
           // -------------------------------------------------------
       10: // Esperar a que el KRC pida número de programa (PGNO_REQ = 1)
           IF #ROB_PGNO_REQ THEN
               // Latch del programa seleccionado (1..3). Forzamos límites por seguridad.
               IF #ProgSel < USINT#1 THEN
                   #pgnoLatched := USINT#1;
               ELSIF #ProgSel > USINT#3 THEN
                   #pgnoLatched := USINT#3;
               ELSE
                   #pgnoLatched := #ProgSel;
               END_IF;

               #step := 20;
           END_IF;


       20: // Presentar PGNO MIENTRAS PGNO_REQ = 1
           IF #ROB_PGNO_REQ THEN
               // Escribir bits binarios 101..108 a partir de #pgnoLatched
               #PGNO_101 := ((#pgnoLatched AND USINT#1) <> USINT#0);
               #PGNO_102 := ((#pgnoLatched AND USINT#2) <> USINT#0);
               #PGNO_103 := ((#pgnoLatched AND USINT#4) <> USINT#0);
               #PGNO_104 := ((#pgnoLatched AND USINT#8) <> USINT#0);
               #PGNO_105 := ((#pgnoLatched AND USINT#16) <> USINT#0);
               #PGNO_106 := ((#pgnoLatched AND USINT#32) <> USINT#0);
               #PGNO_107 := ((#pgnoLatched AND USINT#64) <> USINT#0);
               #PGNO_108 := ((#pgnoLatched AND USINT#128) <> USINT#0);

               // Paridad "even": XOR de los 8 bits (1 si nº de unos es impar)
               #PGNO_PARITY :=
               #PGNO_101 XOR #PGNO_102 XOR #PGNO_103 XOR #PGNO_104 XOR
               #PGNO_105 XOR #PGNO_106 XOR #PGNO_107 XOR #PGNO_108;

               // Arrancamos el TON de estabilidad y pasamos a validación
               #tStable(IN := TRUE,
                        PT := #stableTime);
               #step := 21;
           END_IF;


       21: // Esperar estabilidad y marcar PGNO_VALID
           #tStable(IN := (#step = 21),
                    PT := #stableTime);
           IF #tStable.Q THEN
               #PGNO_VALID := TRUE;        // el KRC ya puede muestrear PGNO
               #step := 22;
           END_IF;


       22: // Mantener PGNO_VALID hasta la CAÍDA de PGNO_REQ
           #PGNO_VALID := TRUE;
           IF #fPgnoReq.Q THEN
               #PGNO_VALID := FALSE;    // cerrar handshake de selección

               // limpiar PGNO para siguientes ciclos
               #PGNO_101 := FALSE;
               #PGNO_102 := FALSE;
               #PGNO_103 := FALSE;
               #PGNO_104 := FALSE;
               #PGNO_105 := FALSE;
               #PGNO_106 := FALSE;
               #PGNO_107 := FALSE;
               #PGNO_108 := FALSE;
               #PGNO_PARITY := FALSE;

               #step := 40;    // → arranque real del programa
           END_IF;

       40: // START real: segundo pulso de $EXT_START para ejecutar el programa
           "ALM_FILTER" := TRUE; // marcador/diagnóstico ELIMINAR
           #tpStart(IN := TRUE,
                    PT := #pulseTime);
           #EXT_START := #tpStart.Q;
           IF NOT #tpStart.Q THEN
               #ROBOT_READY := TRUE;   // handshake completo
               #step := 60;            // → ejecución
           END_IF;


       60: // En ejecución / rearme
           // Para un nuevo ciclo hay que hacer hacer 0→1 de nuevo desde la aplicacion 
           // si #startAutExt no baja, #rStart.Q no volverá a disparar.
           #step := 0;

   END_CASE;
END_REGION
END_FUNCTION_BLOCK

// folder: 20. Robot Services/Mov Manual

FUNCTION_BLOCK "TcpJogging"   // FB5, LAD
{ S7_Optimized_Access := 'TRUE' }
VERSION : 0.1
   VAR_INPUT
      "buttonX+" : Bool;
      "buttonX-" : Bool;
      "buttonY+" : Bool;
      "buttonY-" : Bool;
      "buttonZ+" : Bool;
      "buttonZ-" : Bool;
      "buttonE1+" : Bool;
      "buttonE1-" : Bool;
   END_VAR
BEGIN

REGION Network 1 (SCL): Mapea los valores de los botones de WF
   IF "PlcStatus".mode.effective = 0 THEN

       "Tag_1" := TRUE;
       //MOV X,Y,Z
       //%Q630.0 = buttonX+
       //%Q630.1 = buttonX-
       //%Q630.2 = buttonY+
       //%Q630.3 = buttonY-
       //%Q630.4 = buttonZ+
       //%Q630.5 = buttonZ-
       //MOV A,B,C
       //%Q630.6 = buttonWF +A
       //%Q630.7 = buttonWF -A
       //%Q631.0 = buttonWF +B
       //%Q631.1 = buttonWF -B
       //%Q631.2 = buttonWF +C
       //%Q631.3 = buttonWF -C
       //Mov E1
       //%Q631.4 = buttonWF +E1
       //%Q631.5 = buttonWF -E1

   ELSE
       //%Q631.1 = buttonWF -B
       "Tag_1" := FALSE;
   END_IF;
END_REGION
END_FUNCTION_BLOCK

FUNCTION_BLOCK "TcpTarget"   // FB11, LAD
{ S7_Optimized_Access := 'TRUE' }
VERSION : 0.1
   VAR_INPUT
      KukaControlCmdCode : UInt;
      KukaControlCmdSeq : UInt;
      KukaControlCmdProfileRequestId : UInt;
      KukaControlCmdToolRequestId : UInt;
      KukaControlCmdBaseRequestId : UInt;
      KukaControlCmdProgramRequestId : UInt;
      KukaControlTcpTargetX_mm : LReal;
      KukaControlTcpTargetY_mm : LReal;
      KukaControlTcpTargetZ_mm : LReal;
      kukaControlE1Target_mm : LReal;
      KukaControlCmdCancelGo : Bool;
      KukaControlCmdPauseGo : Bool;
      KukaControlCmdResumeGo : Bool;
      enterService : Bool;
      KukaControlCmdVel : UInt;
      KukaControlCmdIndex : UInt;
      scanPuntoInicialX : LReal;
      scanPuntoInicialY : LReal;
      scanPuntoInicialZ : LReal;
      scanPuntoInicialE1 : LReal;
      scanPuntoFinalX : LReal;
      scanPuntoFinalY : LReal;
      scanPuntoFinalZ : LReal;
      scanPuntoFinalE1 : LReal;
   END_VAR
   VAR_OUTPUT
      moveCodeKuka : Word;
      profileReqId : Word;
      baseReqId : Word;
      toolReqId : Word;
      programReqId : Word;
      x_mmHe : DWord;
      y_mmHe : DWord;
      z_mmHe : DWord;
      e_mmHe : DWord;
      PlcStatusExecDone : Bool;
      PlcStatusExecAccepted : Bool;
      PlcStatusExecAckSeq : UInt;
      PlcStatusExecBusy : Bool;
      PlcStatusExecError : Bool;
      PlcStatusExecErrorCode : DWord;
      PlcStatusExecLastCode : UInt;
      vel_mmsHe : Word;
      index_mmHe : Word;
      xInicial_mm : DWord;
      yInicial_mm : DWord;
      zInicial_mm : DWord;
      e1Inicial_mm : DWord;
      xFinal_mm : DWord;
      yFinal_mm : DWord;
      zFinal_mm : DWord;
      e1Final_mm : DWord;
   END_VAR
   VAR
      lastSeq : UInt;
      lastCode : UInt;
      state : Int;
      tmoMove : TON_TIME;
      rbDoneEdge : R_TRIG;
      _cancelInFlight : Bool := false;   // marca que el DONE que venga es por cancelación
      _isMotion : Bool;   // helper para saber si el code es de movimiento
      rbDoneEdge_1 : R_TRIG;
      rEnterSrv : R_TRIG;
   END_VAR
   VAR_TEMP
      x_dint : DInt;
      y_dint : DInt;
      z_dint : DInt;
      n_dint : DInt;
      code_int : UInt;
      tool_int : UInt;
      xInicial_dint : DInt;
      yInicial_Dint : DInt;
      ZInicial_Dint : DInt;
      e1Inicial_Dint : DInt;
      xFinal_Dint : DInt;
      yFinal_Dint : DInt;
      ZFinal_Dint : DInt;
      e1Final_Dint : DInt;
      index_uint : UInt;
      vel_uint : UInt;
   END_VAR
BEGIN

REGION Network 1 (SCL)
   #rEnterSrv(CLK := #enterService);
   IF #rEnterSrv.Q THEN
       #state := 0;
       #PlcStatusExecAccepted := FALSE;
       #PlcStatusExecBusy := FALSE;
       #PlcStatusExecDone := FALSE;

       // deja lastSeq "uno por detrás" del actual
       IF #KukaControlCmdSeq = UINT#0 THEN
           #lastSeq := UINT#65535;
       ELSE
           #lastSeq := #KukaControlCmdSeq - UINT#1;
       END_IF;
   END_IF;




   CASE #state OF
       0: // IDLE -> GO == ACK
           #PlcStatusExecAccepted := FALSE;
           #PlcStatusExecBusy := FALSE;
           #PlcStatusExecError := FALSE;
           "cancelGo" := FALSE;
           //#PlcStatusExecDone := FALSE;

           #code_int := #KukaControlCmdCode;  // refresca SIEMPRE

           #tool_int := #KukaControlCmdToolRequestId;

           // Nuevo comando si llega seq distinto y el canal está libre
           IF (#KukaControlCmdSeq <> #lastSeq) AND ("goTrigger" = "rbDone") THEN

                   IF #code_int = 130 THEN
                       //  Primero: Escalar mm → entero (µm). Ajusta el redondeo si lo prefieres TRUNC, FLOOR, etc.
                       #n_dint := LREAL_TO_DINT(ROUND(#kukaControlE1Target_mm));
                       // Segundo Convertir a DWORD y hacer SWAP para que el KRC lo lea correctamente
                       #e_mmHe := SWAP(DINT_TO_DWORD(#n_dint));
                   END_IF;

                   IF #code_int = 101 THEN
                       //  Primero: Escalar mm → entero (µm). Ajusta el redondeo si lo prefieres TRUNC, FLOOR, etc.
                       #x_dint := LREAL_TO_DINT(ROUND(#KukaControlTcpTargetX_mm));
                       // Segundo Convertir a DWORD y hacer SWAP para que el KRC lo lea correctamente
                       #x_mmHe := SWAP(DINT_TO_DWORD(#x_dint));
                   END_IF;

                   IF #code_int = 102 THEN
                       //  Primero: Escalar mm → entero (µm). Ajusta el redondeo si lo prefieres TRUNC, FLOOR, etc.
                       #y_dint := LREAL_TO_DINT(ROUND(#KukaControlTcpTargetY_mm));
                       // Segundo Convertir a DWORD y hacer SWAP para que el KRC lo lea correctamente
                       #y_mmHe := SWAP(DINT_TO_DWORD(#y_dint));
                   END_IF;

                   IF #code_int = 103 THEN
                       //  Primero: Escalar mm → entero (µm). Ajusta el redondeo si lo prefieres TRUNC, FLOOR, etc.
                       #z_dint := LREAL_TO_DINT(ROUND(#KukaControlTcpTargetZ_mm));
                       // Segundo Convertir a DWORD y hacer SWAP para que el KRC lo lea correctamente
                       #z_mmHe := SWAP(DINT_TO_DWORD(#z_dint));
                   END_IF;

                   IF #code_int = 201 THEN
                       // id de herramienta → WORD+SWAP
                       #toolReqId := SWAP(UINT_TO_WORD(#KukaControlCmdToolRequestId));

                   END_IF;

                   IF #code_int = 202 THEN

                       // id de herramienta → WORD+SWAP
                       #baseReqId := SWAP(UINT_TO_WORD(#KukaControlCmdBaseRequestId));

                   END_IF;

                   IF #code_int = 203 THEN

                       // id de herramienta → WORD+SWAP
                       #profileReqId := SWAP(UINT_TO_WORD(#KukaControlCmdProfileRequestId));

                   END_IF;

                   // ---------- TEACHING ----------
                   IF #code_int = 301 THEN // Teach Request
                       #programReqId := SWAP(UINT_TO_WORD(#KukaControlCmdProgramRequestId));

                   END_IF;

                   // ---------- TEACH SET START (desde SCA vía OPC) ----------
                   IF #code_int = 311 THEN

                       // Program ID (WORD + SWAP)
                       #programReqId := SWAP(UINT_TO_WORD(#KukaControlCmdProgramRequestId));


                       // Start desde OPC (mm -> DINT -> DWORD + SWAP)
                       //  Primero: Escalar mm → entero (µm). 
                       #xInicial_dint := LREAL_TO_DINT(ROUND(#scanPuntoInicialX));
                       // Segundo Convertir a DWORD y hacer SWAP para que el KRC lo lea correctamente
                       #xInicial_mm := SWAP(DINT_TO_DWORD(#xInicial_dint));
                       #yInicial_Dint := LREAL_TO_DINT(ROUND(#scanPuntoInicialY));
                       #yInicial_mm := SWAP(DINT_TO_DWORD(#yInicial_Dint));
                       #ZInicial_Dint := LREAL_TO_DINT(ROUND(#scanPuntoInicialZ));
                       #zInicial_mm := SWAP(DINT_TO_DWORD(#ZInicial_Dint));
                       #e1Inicial_Dint := LREAL_TO_DINT(ROUND(#scanPuntoInicialE1));
                       #e1Inicial_mm := SWAP(DINT_TO_DWORD(#e1Inicial_Dint));

                   END_IF;

                   // ---------- TEACH SET END (desde SCA vía OPC) ----------
                   IF #code_int = 312 THEN
                       // Program ID también aquí (por robustez)
                       #programReqId := SWAP(UINT_TO_WORD(#KukaControlCmdProgramRequestId));

                       // End desde OPC (mm -> DINT -> DWORD + SWAP)
                       #xFinal_Dint := LREAL_TO_DINT(ROUND(#scanPuntoFinalX));
                       #xFinal_mm := SWAP(DINT_TO_DWORD(#xFinal_Dint));
                       #yFinal_Dint := LREAL_TO_DINT(ROUND(#scanPuntoFinalY));
                       #yFinal_mm := SWAP(DINT_TO_DWORD(#yFinal_Dint));
                       #ZFinal_Dint := LREAL_TO_DINT(ROUND(#scanPuntoFinalZ));
                       #zFinal_mm := SWAP(DINT_TO_DWORD(#ZFinal_Dint));
                       #e1Final_Dint := LREAL_TO_DINT(ROUND(#scanPuntoFinalE1));
                       #e1Final_mm := SWAP(DINT_TO_DWORD(#e1Final_Dint));

                   END_IF;

                   // ---------- SCAN ----------
                   IF #code_int = 402 THEN

                       #programReqId := SWAP(UINT_TO_WORD(#KukaControlCmdProgramRequestId));

                       // ===== START: mm (LREAL) -> DINT -> DWORD + SWAP =====
                       #xInicial_dint := LREAL_TO_DINT(ROUND(#scanPuntoInicialX));
                       #xInicial_mm := SWAP(DINT_TO_DWORD(#xInicial_dint));

                       #yInicial_Dint := LREAL_TO_DINT(ROUND(#scanPuntoInicialY));
                       #yInicial_mm := SWAP(DINT_TO_DWORD(#yInicial_Dint));

                       #ZInicial_Dint := LREAL_TO_DINT(ROUND(#scanPuntoInicialZ));
                       #zInicial_mm := SWAP(DINT_TO_DWORD(#ZInicial_Dint));

                       #e1Inicial_Dint := LREAL_TO_DINT(ROUND(#scanPuntoInicialE1));
                       #e1Inicial_mm := SWAP(DINT_TO_DWORD(#e1Inicial_Dint));

                       // ===== END: mm (LREAL) -> DINT -> DWORD + SWAP =====
                       #xFinal_Dint := LREAL_TO_DINT(ROUND(#scanPuntoFinalX));
                       #xFinal_mm := SWAP(DINT_TO_DWORD(#xFinal_Dint));

                       #yFinal_Dint := LREAL_TO_DINT(ROUND(#scanPuntoFinalY));
                       #yFinal_mm := SWAP(DINT_TO_DWORD(#yFinal_Dint));

                       #ZFinal_Dint := LREAL_TO_DINT(ROUND(#scanPuntoFinalZ));
                       #zFinal_mm := SWAP(DINT_TO_DWORD(#ZFinal_Dint));

                       #e1Final_Dint := LREAL_TO_DINT(ROUND(#scanPuntoFinalE1));
                       #e1Final_mm := SWAP(DINT_TO_DWORD(#e1Final_Dint));

                       // ===== Opcional pero recomendado: velocidad e índice =====
                       // Si en KRC tienes mapeadas variables para vel/index:
                       #vel_uint := #KukaControlCmdVel;
                       #index_uint := #KukaControlCmdIndex;
                       #vel_mmsHe := SWAP(UINT_TO_WORD(#vel_uint));
                       #index_mmHe := SWAP(UINT_TO_WORD(#index_uint));
                       // #index_Dint  := LREAL_TO_DINT(ROUND(#KukaControlCmd_index_mm));
                       // #index_mmHe  := SWAP(DINT_TO_DWORD(#index_Dint));

                   END_IF;



                   // Segundo Convertir a DWORD y hacer SWAP para que el KRC lo lea correctamente
                   #moveCodeKuka := SWAP(UINT_TO_WORD(#code_int));
                   // "moveCodeKuka" := SWAP(UINT_TO_WORD(#code_int));

                   // Dispara GO (flanco por nivel)
                   "goTrigger" := NOT "goTrigger";     // Dispara pedido

                   // Marca estado/ack interno
                   #PlcStatusExecAccepted := TRUE;
                   #PlcStatusExecBusy := TRUE;
                   #PlcStatusExecDone := FALSE;

                   #lastSeq := #KukaControlCmdSeq;          // <-- memoriza!
                   #lastCode := #code_int;             // memoriza qué comando es (para actualizar activos en DONE)

                   #state := 20;                    // BUSY


       END_IF;

   20: // BUSY

       #PlcStatusExecBusy := TRUE;

       #code_int := #KukaControlCmdCode;

       // CANCEL pedido en BUSY → avisar al KRC y ACK de la ORDEN ACTIVA
       IF #code_int = 903 THEN
           "cancelGo" := TRUE;
       END_IF;

       IF ("rbDone" = "goTrigger") THEN
           // Fin confirmado por KUKA

           #PlcStatusExecDone := TRUE;
           #PlcStatusExecBusy := FALSE;
           #PlcStatusExecAccepted := FALSE;
           // ACK de la orden completada
           #PlcStatusExecAckSeq := #lastSeq;

           #state := 0;                         // vuelve a IDLE

       END_IF;

   30: // DONE
       // limpiar y volver a IDLE
       #state := 0;


   END_CASE;
END_REGION
END_FUNCTION_BLOCK

// folder: 20. Robot Services/RobotPos

FUNCTION_BLOCK "TcpPoseDecoderLe32"   // FB4, LAD
{ S7_Optimized_Access := 'TRUE' }
VERSION : 0.1
// Decodifica con SWAP, convierte a DINT y escala.
   VAR_INPUT
      xIniRawLe : DWord;
      yIniRawLe : DWord;
      zIniRawLe : DWord;
      e1IniRawLe : DWord;
      xFinRawLe : DWord;
      yFinRawLe : DWord;
      zFinRawLe : DWord;
      e1FinRawLe : DWord;
      ToolActiveRawByte : Byte;
      BaseActiveRawByte : Byte;
   END_VAR
   VAR_OUTPUT
      tcpPosIniX_mm : LReal;
      tcpPosIniY_mm : LReal;
      tcpPosIniZ_mm : LReal;
      e1PosIni_mm : LReal;
      tcpPosFinX_mm : LReal;
      tcpPosFinY_mm : LReal;
      tcpPosFinZ_mm : LReal;
      e1PosFin_mm : LReal;
      toolActiveId : UDInt;
      baseActiveId : UDInt;
   END_VAR
   VAR_TEMP
      xIniDint : DInt;
      yIniDint : DInt;
      zIniDint : DInt;
      aDint : DInt;
      bDint : DInt;
      cDint : DInt;
      e1IniDint : DInt;
      xFinDint : DInt;
      yFinDint : DInt;
      zFinDint : DInt;
      e1FinDint : DInt;
   END_VAR
BEGIN

REGION Network 1 (SCL): // 1) Endianness: ABCD -> DCBA
   #xIniDint := DWORD_TO_DINT(SWAP(#xIniRawLe));
   #yIniDint := DWORD_TO_DINT(SWAP(#yIniRawLe));
   #zIniDint := DWORD_TO_DINT(SWAP(#zIniRawLe));

   #e1IniDint := DWORD_TO_DINT(SWAP(#e1IniRawLe));

   #xFinDint := DWORD_TO_DINT(SWAP(#xFinRawLe));
   #yFinDint := DWORD_TO_DINT(SWAP(#yFinRawLe));
   #zFinDint := DWORD_TO_DINT(SWAP(#zFinRawLe));
   #e1FinDint := DWORD_TO_DINT(SWAP(#e1FinRawLe));
END_REGION

REGION Network 2 (SCL): // 2) Escala fixed-point: µm->mm, mdeg->deg
   #tcpPosIniX_mm := DINT_TO_LREAL(#xIniDint) / 1000.0;
   #tcpPosIniY_mm := DINT_TO_LREAL(#yIniDint) / 1000.0;
   #tcpPosIniZ_mm := DINT_TO_LREAL(#zIniDint) / 1000.0;

   #e1PosIni_mm := DINT_TO_LREAL(#e1IniDint) / 1000.0;  // mm o deg según tu E1

   #tcpPosFinX_mm := DINT_TO_LREAL(#xFinDint) / 1000.0;
   #tcpPosFinY_mm := DINT_TO_LREAL(#yFinDint) / 1000.0;
   #tcpPosFinZ_mm := DINT_TO_LREAL(#zFinDint) / 1000.0;
   #e1PosFin_mm := DINT_TO_LREAL(#e1FinDint) / 1000.0;  // mm o deg según tu E1

   #toolActiveId := #ToolActiveRawByte;
   #baseActiveId := #BaseActiveRawByte;
END_REGION
END_FUNCTION_BLOCK

// folder: 20. Robot Services/Tooling & Parking

FUNCTION_BLOCK "ToolChange"   // FB6, LAD
TITLE = FB: ManageTed009Station
{ S7_Optimized_Access := 'TRUE' }
VERSION : 0.1
// //  - KUKA manda órdenes (kukaCmd*)
// //  - El FB acciona bobinas de la docking (dockValve*On)
// //  - El FB publica ecos/estados para el KUKA (kukaFeedback*)
// //  - V2 (Unlock) puede mantenerse automática con útil aparcado
// //    (AutoUnlockWhenToolPresent = TRUE) [REF: estándar automático]. 
// //    Con útil ausente, no se activa para evitar soplado innecesario.
// //  - Tapa: FSM con interlock de zona segura y timeouts simétricos.
// //  - Diagnóstico: diagStep/diagFault/diagFaultCode.
// //
// //  Referencias (ver manual Stäubli TED009):
// //    • Sequence plan y sondeo ~20 ms durante conectar/desconectar. 
// //    • +21 mm: E2=0 ∧ E3=1 ∧ D1=0 antes de acoplar. 
// //    • z=0: bloquear retirando V2 y esperar E2=1 ∧ D1=1 (+E1=1). 
// //    • Retiradas +10/+70 y +25/>29 (comentadas para el programa del robot).
   VAR_INPUT
      kukaCmdOpenCover : Bool;
      kukaCmdCloseCover : Bool;
      kukaCmdUnlockMps : Bool;
      kukaCmdSafeForChange : Bool;
      dockSensorToolInPosition : Bool;   // E6
      dockSensorCoverClosed : Bool;   // E4
      dockSensorCoverOpen : Bool;   // E5
      robotSensorMpsUnlocked : Bool;   // E3
      robotSensorMpsLocked : Bool;   // E2
      robotSensorMpsCoupled : Bool;   // E1
      robotSensorMpsCtrlAirPressureOk : Bool;   // D1
      resetFault : Bool;
   END_VAR
   VAR_OUTPUT
      dockValveCoverOpenOn : Bool;   // bobina abrir tapa
      dockValveCoverCloseOn : Bool;   // bobina cerrar tapa
      dockValveV2UnlockOn : Bool;   // V2: aire de desbloqueo hacia módulo del robot
      MpsValveV1B12S4_ON : Bool;
      kukaFeedbackDockCoverOpen : Bool;
      kukaFeedbackDockCoverClosed : Bool;
      kukaFeedbackRobotMpsUnlocked : Bool;
      kukaFeedbackRobotMpsLocked : Bool;
      kukaFeedbackRobotMpsCoupled : Bool;
      kukaFeedbackMpsCtrlAirPressureOk : Bool;
      kukaFeedbackDockToolInPosition : Bool;
      diagStep : Int;
      diagFault : Bool;
      diagFaultCode : Int;
   END_VAR
   VAR
      "step" : Int;
      fault : Bool;
      faultCode : Int;
      AutoUnlockWhenToolPresent : Bool := true;   // // modo auto
      coverTimeout : Time := T#8S;   // // timeout de tapa (abrir/cerrar)
      unlockTimeout : Time := T#2S;   // // timeout de UNLOCK (E3=1 & D1=0)
      unlockReq : Bool;
      unlockReqEnabled : Bool;
      tempCoverOpen : TON_TIME;
      tempCoverClose : TON_TIME;
      tempUnlock : TON_TIME;
      autoUnlockEligible : Bool;
   END_VAR
   VAR CONSTANT
      StateIdle : Int := 0;
      StateOpening : Int := 10;
      StateOpen : Int := 11;
      StateClosing : Int := 20;
      StateClosed : Int := 21;
      FaultNone : Int;
      FaultOpenTimeout : Int := 101;
      FaultCloseTimeout : Int := 102;
      FaultUnlockTimeout : Int := 201;
      FaultInterlock : Int := 301;
   END_VAR
BEGIN

REGION Network 1 (SCL): Lógica de tapa + V2 (Unlock) de la docking
   // --- Feedbacks de estados al robot (eco directo de sensores físicos)
   #kukaFeedbackDockToolInPosition := #dockSensorToolInPosition; // E6 - herramienta en docking station
   #kukaFeedbackDockCoverOpen := #dockSensorCoverOpen;         // E4 - tapa abierta
   #kukaFeedbackDockCoverClosed := #dockSensorCoverClosed;     // E5 - tapa cerrada
   #kukaFeedbackRobotMpsUnlocked := #robotSensorMpsUnlocked;  // E3 - MPS desbloqueado (robot side)
   #kukaFeedbackRobotMpsLocked := #robotSensorMpsLocked;     // E2 - MPS bloqueado (robot side
   #kukaFeedbackRobotMpsCoupled := #robotSensorMpsCoupled;        // E1 - MPS acoplado  (robot side) 
   #kukaFeedbackMpsCtrlAirPressureOk := #robotSensorMpsCtrlAirPressureOk;  // D1 -presostato módulo aire control (robot)
   // ---- Reset de fallos/estado -------------------------------------------
   // Permite reconocer fallos desde HMI/Robot. Pone las salidas a 0 y la FSM (flow state machine)
   // Deja el FB en reposo (IDLE), corta bobinas y reinicia tempor TONs.
   // 
   IF #resetFault THEN
       #fault := FALSE;
       #faultCode := #FaultNone;
       #step := #StateIdle;

       #dockValveCoverOpenOn := FALSE;
       #dockValveCoverCloseOn := FALSE;
       #dockValveV2UnlockOn := FALSE;

       // Reset explícito de TON: IN=FALSE + PT definido
       #tempCoverOpen(IN := FALSE,
                      PT := #coverTimeout);
       #tempCoverClose(IN := FALSE,
                       PT := #coverTimeout);
       #tempUnlock(IN := FALSE,
                   PT := #unlockTimeout);
   END_IF;

   // ================= LÓGICA DE TAPA (máquina de estados) =================
   // Interlock básico: no se permite accionar tapa si el robot no confirma zona segura
   // (manual: abrir/cerrar solo fuera del barrido).
   CASE #step OF

       #StateIdle: // IDLE
           // Reposo ( tapa sin accionar); evaluar órdenes de KUKA.
           #dockValveCoverOpenOn := FALSE;
           #dockValveCoverCloseOn := FALSE;

           IF #kukaCmdSafeForChange THEN
               // Abrir si lo pide el robot y aún no está abierta
               IF (#kukaCmdOpenCover AND NOT #dockSensorCoverOpen) THEN
                   #step := #StateOpening;
               END_IF;
               // Cerrar si lo pide el robot y aún no está cerrada
               IF (#kukaCmdCloseCover AND NOT #dockSensorCoverClosed) THEN
                   #step := #StateClosing;
               END_IF;
           ELSIF (#kukaCmdOpenCover OR #kukaCmdCloseCover) THEN
               // Petición sin zona segura -> fallo de interlock
               #fault := TRUE;
               #faultCode := #FaultInterlock; // robot no garantiza zona segura
           END_IF;

       #StateOpening:  // Abrir tapa
           #dockValveCoverOpenOn := TRUE;
           #dockValveCoverCloseOn := FALSE;

           // Timeout de apertura: si no llega "tapa abierta" dentro de coverTimeout -> fallo.
           // coverTimeout debe ser > 3 s (tiempo típico de maniobra)
           #tempCoverOpen(IN := NOT #dockSensorCoverOpen,
                          PT := #coverTimeout);

           IF (#dockSensorCoverOpen AND NOT #dockSensorCoverClosed) THEN
               #tempCoverOpen(IN := FALSE,
                              PT := #coverTimeout);
               #step := #StateOpen;
           ELSIF #tempCoverOpen.Q THEN
               #fault := TRUE;
               #faultCode := #FaultOpenTimeout;
               #dockValveCoverOpenOn := FALSE;
               #step := #StateIdle;
           END_IF;

       #StateOpen: // Tapa abierta (estable)
           #dockValveCoverOpenOn := FALSE;
           #dockValveCoverCloseOn := FALSE;

           IF (#kukaCmdSafeForChange AND #kukaCmdCloseCover) THEN
               #step := #StateClosing;
           END_IF;


       #StateClosing: // Cerrar tapa
           #dockValveCoverOpenOn := FALSE;
           #dockValveCoverCloseOn := TRUE;

           // Timeout de cierre: si no llega "tapa cerrada" dentro de coverTimeout -> fallo.
           #tempCoverClose(IN := NOT #dockSensorCoverClosed,
                           PT := #coverTimeout);

           IF (#dockSensorCoverClosed AND NOT #dockSensorCoverOpen) THEN
               #tempCoverClose(IN := FALSE,
                               PT := #coverTimeout);
               #step := #StateClosed;
           ELSIF #tempCoverClose.Q THEN
               #fault := TRUE;
               #faultCode := #FaultCloseTimeout;
               #dockValveCoverCloseOn := FALSE;
               #step := #StateIdle;
           END_IF;

       #StateClosed: // Tapa cerrada (estable)
           #dockValveCoverOpenOn := FALSE;
           #dockValveCoverCloseOn := FALSE;

           IF (#kukaCmdSafeForChange AND #kukaCmdOpenCover) THEN
               #step := #StateOpening;
           END_IF;

       ELSE
           #step := #StateIdle;
   END_CASE;

   // Exclusión mutua de bobinas de tapa (seguridad por si alguna rama dejó ambas a 1)
   IF #dockValveCoverOpenOn THEN
       #dockValveCoverCloseOn := FALSE;
   END_IF;
   IF #dockValveCoverCloseOn THEN
       #dockValveCoverOpenOn := FALSE;
   END_IF;



   // -------- Arbitraje de V2 (UNLOCK) — sin auto-unlock --------
   #autoUnlockEligible := FALSE;   // DEPRECATED: ya no se usa

   //Cuando el robot va al punto de acople hace antes kukaCmdUnlockMpsYugo = TRUE

   //  solo por orden KUKA 
   #dockValveV2UnlockOn := #kukaCmdUnlockMps;

   IF #robotSensorMpsLocked THEN
       #MpsValveV1B12S4_ON := TRUE;
   END_IF;


   // Supervisión del estado desbloqueado (E3=1 y D1=0 en tiempo):
   #tempUnlock(
               IN := (#dockValveV2UnlockOn
               AND NOT (#robotSensorMpsUnlocked
               AND NOT #robotSensorMpsCtrlAirPressureOk)),
               PT := #unlockTimeout
   );
   IF NOT #dockValveV2UnlockOn THEN
       // reset explícito del TON cuando ya no se pide V2
       #tempUnlock(IN := FALSE,
                   PT := #unlockTimeout);
   END_IF;

   // -------------------- DIAGNÓSTICO PUBLICADO ----------------------------
   #diagStep := #step; // StateIdle/Opening/Open/Closing/Closed
   #diagFault := #fault;
   #diagFaultCode := #faultCode;
END_REGION
END_FUNCTION_BLOCK

FUNCTION_BLOCK "MpsDockingStation"   // FB9, LAD
{ S7_Optimized_Access := 'TRUE' }
VERSION : 0.1
BEGIN

REGION Network 1: Identificador de Herramienta
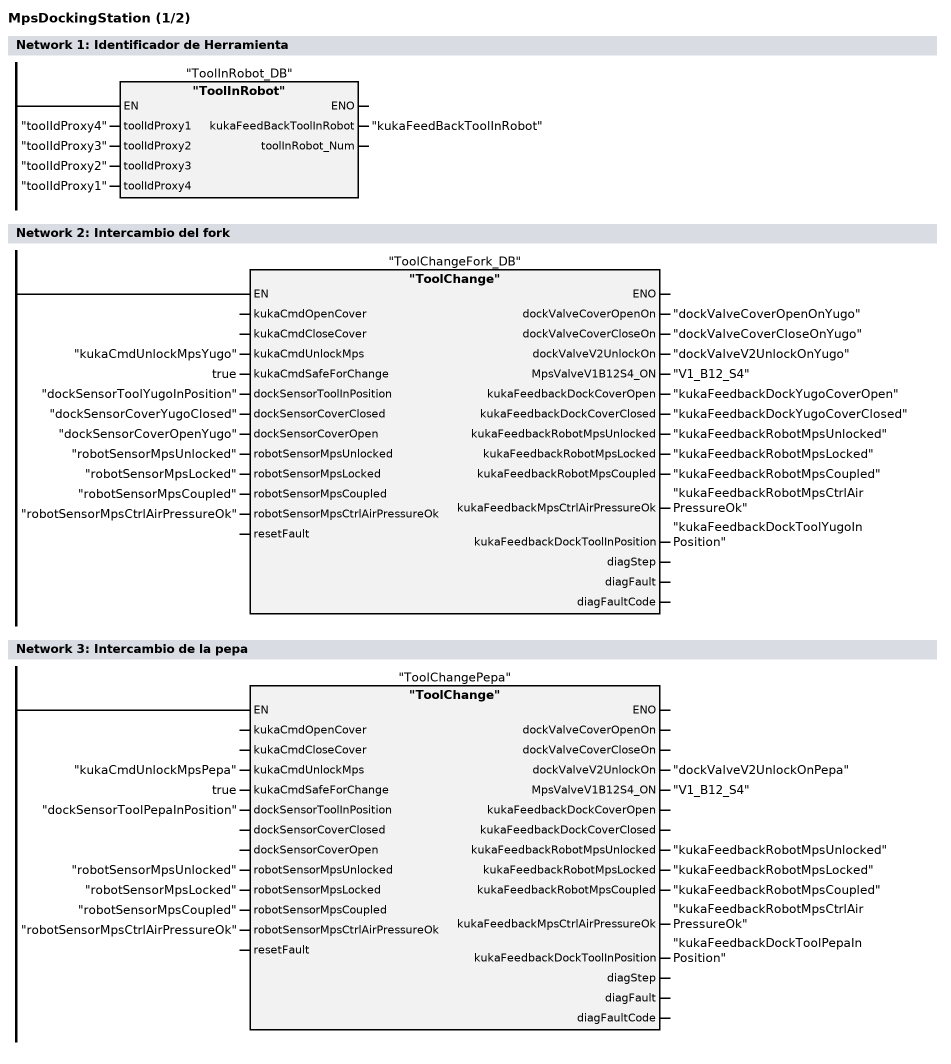
   RUNG wire#powerrail
      "ToolInRobot_DB"(toolIdProxy1 := "toolIdProxy4", toolIdProxy2 := "toolIdProxy3", toolIdProxy3 := "toolIdProxy2", toolIdProxy4 := "toolIdProxy1", kukaFeedBackToolInRobot => "kukaFeedBackToolInRobot", toolInRobot_Num =>)
   END_RUNG
   // the same network as SCL:
   "ToolInRobot_DB"(toolIdProxy1 := "toolIdProxy4",   // "ToolInRobot"
                    toolIdProxy2 := "toolIdProxy3",
                    toolIdProxy3 := "toolIdProxy2",
                    toolIdProxy4 := "toolIdProxy1",
                    kukaFeedBackToolInRobot => "kukaFeedBackToolInRobot");
END_REGION

REGION Network 2: Intercambio del fork
   RUNG wire#powerrail
      "ToolChangeFork_DB"(kukaCmdOpenCover :=, kukaCmdCloseCover :=, kukaCmdUnlockMps := "kukaCmdUnlockMpsYugo", kukaCmdSafeForChange := true, dockSensorToolInPosition := "dockSensorToolYugoInPosition", dockSensorCoverClosed := "dockSensorCoverYugoClosed", dockSensorCoverOpen := "dockSensorCoverOpenYugo", robotSensorMpsUnlocked := "robotSensorMpsUnlocked", robotSensorMpsLocked := "robotSensorMpsLocked", robotSensorMpsCoupled := "robotSensorMpsCoupled", robotSensorMpsCtrlAirPressureOk := "robotSensorMpsCtrlAirPressureOk", resetFault :=, dockValveCoverOpenOn => "dockValveCoverOpenOnYugo", dockValveCoverCloseOn => "dockValveCoverCloseOnYugo", dockValveV2UnlockOn => "dockValveV2UnlockOnYugo", MpsValveV1B12S4_ON => "V1_B12_S4", kukaFeedbackDockCoverOpen => "kukaFeedbackDockYugoCoverOpen", kukaFeedbackDockCoverClosed => "kukaFeedbackDockYugoCoverClosed", kukaFeedbackRobotMpsUnlocked => "kukaFeedbackRobotMpsUnlocked", kukaFeedbackRobotMpsLocked => "kukaFeedbackRobotMpsLocked", kukaFeedbackRobotMpsCoupled => "kukaFeedbackRobotMpsCoupled", kukaFeedbackMpsCtrlAirPressureOk => "kukaFeedbackRobotMpsCtrlAirPressureOk", kukaFeedbackDockToolInPosition => "kukaFeedbackDockToolYugoInPosition", diagStep =>, diagFault =>, diagFaultCode =>)
   END_RUNG
   // the same network as SCL:
   "ToolChangeFork_DB"(kukaCmdUnlockMps := "kukaCmdUnlockMpsYugo",   // "ToolChange"
                       kukaCmdSafeForChange := true,
                       dockSensorToolInPosition := "dockSensorToolYugoInPosition",
                       dockSensorCoverClosed := "dockSensorCoverYugoClosed",
                       dockSensorCoverOpen := "dockSensorCoverOpenYugo",
                       robotSensorMpsUnlocked := "robotSensorMpsUnlocked",
                       robotSensorMpsLocked := "robotSensorMpsLocked",
                       robotSensorMpsCoupled := "robotSensorMpsCoupled",
                       robotSensorMpsCtrlAirPressureOk := "robotSensorMpsCtrlAirPressureOk",
                       dockValveCoverOpenOn => "dockValveCoverOpenOnYugo",
                       dockValveCoverCloseOn => "dockValveCoverCloseOnYugo",
                       dockValveV2UnlockOn => "dockValveV2UnlockOnYugo",
                       MpsValveV1B12S4_ON => "V1_B12_S4",
                       kukaFeedbackDockCoverOpen => "kukaFeedbackDockYugoCoverOpen",
                       kukaFeedbackDockCoverClosed => "kukaFeedbackDockYugoCoverClosed",
                       kukaFeedbackRobotMpsUnlocked => "kukaFeedbackRobotMpsUnlocked",
                       kukaFeedbackRobotMpsLocked => "kukaFeedbackRobotMpsLocked",
                       kukaFeedbackRobotMpsCoupled => "kukaFeedbackRobotMpsCoupled",
                       kukaFeedbackMpsCtrlAirPressureOk => "kukaFeedbackRobotMpsCtrlAirPressureOk",
                       kukaFeedbackDockToolInPosition => "kukaFeedbackDockToolYugoInPosition");
END_REGION

REGION Network 3: Intercambio de la pepa
   RUNG wire#powerrail
      "ToolChangePepa"(kukaCmdOpenCover :=, kukaCmdCloseCover :=, kukaCmdUnlockMps := "kukaCmdUnlockMpsPepa", kukaCmdSafeForChange := true, dockSensorToolInPosition := "dockSensorToolPepaInPosition", dockSensorCoverClosed :=, dockSensorCoverOpen :=, robotSensorMpsUnlocked := "robotSensorMpsUnlocked", robotSensorMpsLocked := "robotSensorMpsLocked", robotSensorMpsCoupled := "robotSensorMpsCoupled", robotSensorMpsCtrlAirPressureOk := "robotSensorMpsCtrlAirPressureOk", resetFault :=, dockValveCoverOpenOn =>, dockValveCoverCloseOn =>, dockValveV2UnlockOn => "dockValveV2UnlockOnPepa", MpsValveV1B12S4_ON => "V1_B12_S4", kukaFeedbackDockCoverOpen =>, kukaFeedbackDockCoverClosed =>, kukaFeedbackRobotMpsUnlocked => "kukaFeedbackRobotMpsUnlocked", kukaFeedbackRobotMpsLocked => "kukaFeedbackRobotMpsLocked", kukaFeedbackRobotMpsCoupled => "kukaFeedbackRobotMpsCoupled", kukaFeedbackMpsCtrlAirPressureOk => "kukaFeedbackRobotMpsCtrlAirPressureOk", kukaFeedbackDockToolInPosition => "kukaFeedbackDockToolPepaInPosition", diagStep =>, diagFault =>, diagFaultCode =>)
   END_RUNG
   // the same network as SCL:
   "ToolChangePepa"(kukaCmdUnlockMps := "kukaCmdUnlockMpsPepa",   // "ToolChange"
                    kukaCmdSafeForChange := true,
                    dockSensorToolInPosition := "dockSensorToolPepaInPosition",
                    robotSensorMpsUnlocked := "robotSensorMpsUnlocked",
                    robotSensorMpsLocked := "robotSensorMpsLocked",
                    robotSensorMpsCoupled := "robotSensorMpsCoupled",
                    robotSensorMpsCtrlAirPressureOk := "robotSensorMpsCtrlAirPressureOk",
                    dockValveV2UnlockOn => "dockValveV2UnlockOnPepa",
                    MpsValveV1B12S4_ON => "V1_B12_S4",
                    kukaFeedbackRobotMpsUnlocked => "kukaFeedbackRobotMpsUnlocked",
                    kukaFeedbackRobotMpsLocked => "kukaFeedbackRobotMpsLocked",
                    kukaFeedbackRobotMpsCoupled => "kukaFeedbackRobotMpsCoupled",
                    kukaFeedbackMpsCtrlAirPressureOk => "kukaFeedbackRobotMpsCtrlAirPressureOk",
                    kukaFeedbackDockToolInPosition => "kukaFeedbackDockToolPepaInPosition");
END_REGION

REGION Network 4: Intercambio de la heramienta de Inmersion - Pole
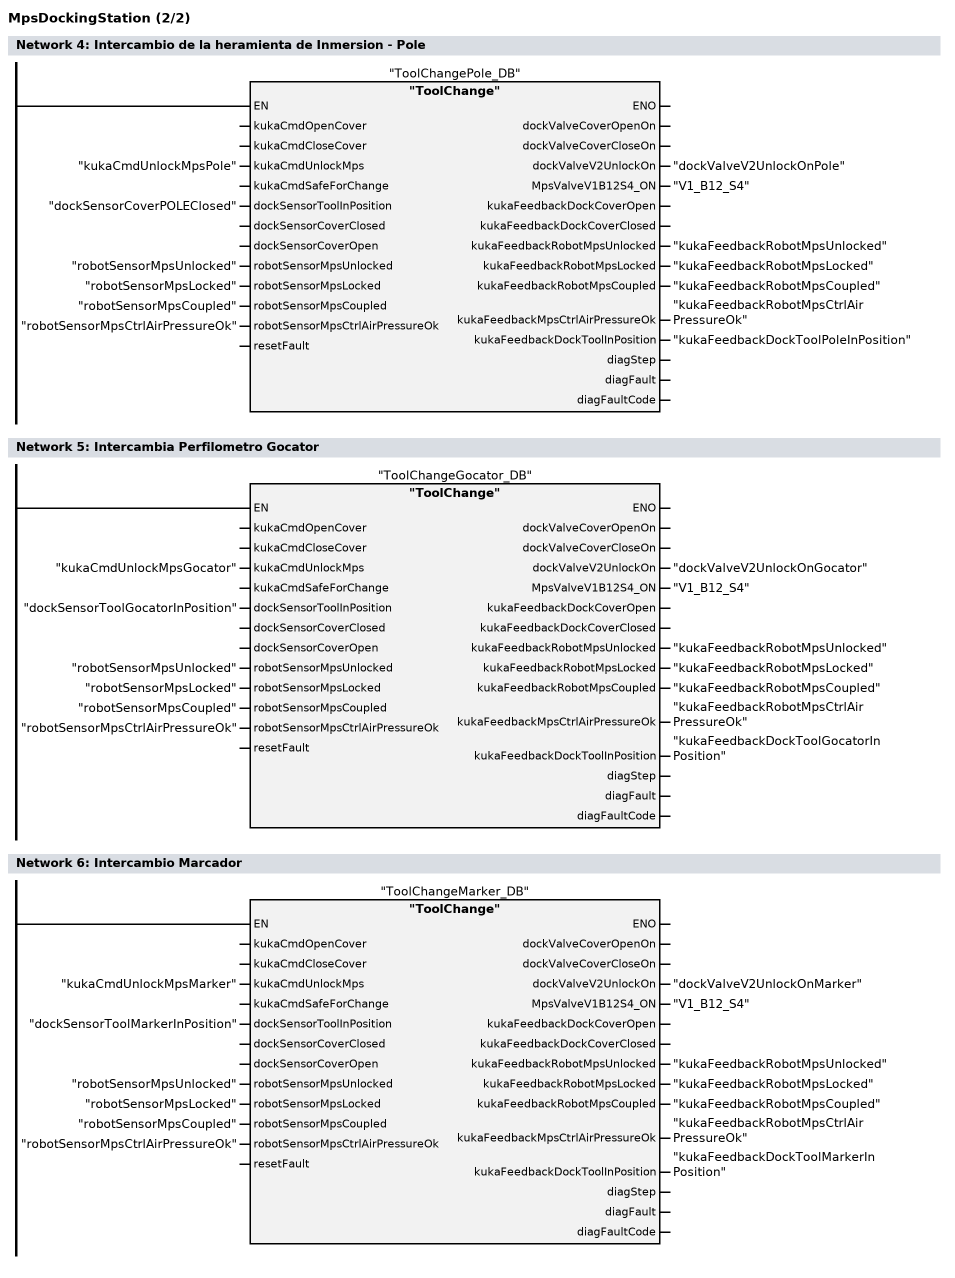
   RUNG wire#powerrail
      "ToolChangePole_DB"(kukaCmdOpenCover :=, kukaCmdCloseCover :=, kukaCmdUnlockMps := "kukaCmdUnlockMpsPole", kukaCmdSafeForChange :=, dockSensorToolInPosition := "dockSensorCoverPOLEClosed", dockSensorCoverClosed :=, dockSensorCoverOpen :=, robotSensorMpsUnlocked := "robotSensorMpsUnlocked", robotSensorMpsLocked := "robotSensorMpsLocked", robotSensorMpsCoupled := "robotSensorMpsCoupled", robotSensorMpsCtrlAirPressureOk := "robotSensorMpsCtrlAirPressureOk", resetFault :=, dockValveCoverOpenOn =>, dockValveCoverCloseOn =>, dockValveV2UnlockOn => "dockValveV2UnlockOnPole", MpsValveV1B12S4_ON => "V1_B12_S4", kukaFeedbackDockCoverOpen =>, kukaFeedbackDockCoverClosed =>, kukaFeedbackRobotMpsUnlocked => "kukaFeedbackRobotMpsUnlocked", kukaFeedbackRobotMpsLocked => "kukaFeedbackRobotMpsLocked", kukaFeedbackRobotMpsCoupled => "kukaFeedbackRobotMpsCoupled", kukaFeedbackMpsCtrlAirPressureOk => "kukaFeedbackRobotMpsCtrlAirPressureOk", kukaFeedbackDockToolInPosition => "kukaFeedbackDockToolPoleInPosition", diagStep =>, diagFault =>, diagFaultCode =>)
   END_RUNG
   // the same network as SCL:
   "ToolChangePole_DB"(kukaCmdUnlockMps := "kukaCmdUnlockMpsPole",   // "ToolChange"
                       dockSensorToolInPosition := "dockSensorCoverPOLEClosed",
                       robotSensorMpsUnlocked := "robotSensorMpsUnlocked",
                       robotSensorMpsLocked := "robotSensorMpsLocked",
                       robotSensorMpsCoupled := "robotSensorMpsCoupled",
                       robotSensorMpsCtrlAirPressureOk := "robotSensorMpsCtrlAirPressureOk",
                       dockValveV2UnlockOn => "dockValveV2UnlockOnPole",
                       MpsValveV1B12S4_ON => "V1_B12_S4",
                       kukaFeedbackRobotMpsUnlocked => "kukaFeedbackRobotMpsUnlocked",
                       kukaFeedbackRobotMpsLocked => "kukaFeedbackRobotMpsLocked",
                       kukaFeedbackRobotMpsCoupled => "kukaFeedbackRobotMpsCoupled",
                       kukaFeedbackMpsCtrlAirPressureOk => "kukaFeedbackRobotMpsCtrlAirPressureOk",
                       kukaFeedbackDockToolInPosition => "kukaFeedbackDockToolPoleInPosition");
END_REGION

REGION Network 5: Intercambia Perfilometro Gocator
   RUNG wire#powerrail
      "ToolChangeGocator_DB"(kukaCmdOpenCover :=, kukaCmdCloseCover :=, kukaCmdUnlockMps := "kukaCmdUnlockMpsGocator", kukaCmdSafeForChange :=, dockSensorToolInPosition := "dockSensorToolGocatorInPosition", dockSensorCoverClosed :=, dockSensorCoverOpen :=, robotSensorMpsUnlocked := "robotSensorMpsUnlocked", robotSensorMpsLocked := "robotSensorMpsLocked", robotSensorMpsCoupled := "robotSensorMpsCoupled", robotSensorMpsCtrlAirPressureOk := "robotSensorMpsCtrlAirPressureOk", resetFault :=, dockValveCoverOpenOn =>, dockValveCoverCloseOn =>, dockValveV2UnlockOn => "dockValveV2UnlockOnGocator", MpsValveV1B12S4_ON => "V1_B12_S4", kukaFeedbackDockCoverOpen =>, kukaFeedbackDockCoverClosed =>, kukaFeedbackRobotMpsUnlocked => "kukaFeedbackRobotMpsUnlocked", kukaFeedbackRobotMpsLocked => "kukaFeedbackRobotMpsLocked", kukaFeedbackRobotMpsCoupled => "kukaFeedbackRobotMpsCoupled", kukaFeedbackMpsCtrlAirPressureOk => "kukaFeedbackRobotMpsCtrlAirPressureOk", kukaFeedbackDockToolInPosition => "kukaFeedbackDockToolGocatorInPosition", diagStep =>, diagFault =>, diagFaultCode =>)
   END_RUNG
   // the same network as SCL:
   "ToolChangeGocator_DB"(kukaCmdUnlockMps := "kukaCmdUnlockMpsGocator",   // "ToolChange"
                          dockSensorToolInPosition := "dockSensorToolGocatorInPosition",
                          robotSensorMpsUnlocked := "robotSensorMpsUnlocked",
                          robotSensorMpsLocked := "robotSensorMpsLocked",
                          robotSensorMpsCoupled := "robotSensorMpsCoupled",
                          robotSensorMpsCtrlAirPressureOk := "robotSensorMpsCtrlAirPressureOk",
                          dockValveV2UnlockOn => "dockValveV2UnlockOnGocator",
                          MpsValveV1B12S4_ON => "V1_B12_S4",
                          kukaFeedbackRobotMpsUnlocked => "kukaFeedbackRobotMpsUnlocked",
                          kukaFeedbackRobotMpsLocked => "kukaFeedbackRobotMpsLocked",
                          kukaFeedbackRobotMpsCoupled => "kukaFeedbackRobotMpsCoupled",
                          kukaFeedbackMpsCtrlAirPressureOk => "kukaFeedbackRobotMpsCtrlAirPressureOk",
                          kukaFeedbackDockToolInPosition => "kukaFeedbackDockToolGocatorInPosition");
END_REGION

REGION Network 6: Intercambio Marcador
   RUNG wire#powerrail
      "ToolChangeMarker_DB"(kukaCmdOpenCover :=, kukaCmdCloseCover :=, kukaCmdUnlockMps := "kukaCmdUnlockMpsMarker", kukaCmdSafeForChange :=, dockSensorToolInPosition := "dockSensorToolMarkerInPosition", dockSensorCoverClosed :=, dockSensorCoverOpen :=, robotSensorMpsUnlocked := "robotSensorMpsUnlocked", robotSensorMpsLocked := "robotSensorMpsLocked", robotSensorMpsCoupled := "robotSensorMpsCoupled", robotSensorMpsCtrlAirPressureOk := "robotSensorMpsCtrlAirPressureOk", resetFault :=, dockValveCoverOpenOn =>, dockValveCoverCloseOn =>, dockValveV2UnlockOn => "dockValveV2UnlockOnMarker", MpsValveV1B12S4_ON => "V1_B12_S4", kukaFeedbackDockCoverOpen =>, kukaFeedbackDockCoverClosed =>, kukaFeedbackRobotMpsUnlocked => "kukaFeedbackRobotMpsUnlocked", kukaFeedbackRobotMpsLocked => "kukaFeedbackRobotMpsLocked", kukaFeedbackRobotMpsCoupled => "kukaFeedbackRobotMpsCoupled", kukaFeedbackMpsCtrlAirPressureOk => "kukaFeedbackRobotMpsCtrlAirPressureOk", kukaFeedbackDockToolInPosition => "kukaFeedbackDockToolMarkerInPosition", diagStep =>, diagFault =>, diagFaultCode =>)
   END_RUNG
   // the same network as SCL:
   "ToolChangeMarker_DB"(kukaCmdUnlockMps := "kukaCmdUnlockMpsMarker",   // "ToolChange"
                         dockSensorToolInPosition := "dockSensorToolMarkerInPosition",
                         robotSensorMpsUnlocked := "robotSensorMpsUnlocked",
                         robotSensorMpsLocked := "robotSensorMpsLocked",
                         robotSensorMpsCoupled := "robotSensorMpsCoupled",
                         robotSensorMpsCtrlAirPressureOk := "robotSensorMpsCtrlAirPressureOk",
                         dockValveV2UnlockOn => "dockValveV2UnlockOnMarker",
                         MpsValveV1B12S4_ON => "V1_B12_S4",
                         kukaFeedbackRobotMpsUnlocked => "kukaFeedbackRobotMpsUnlocked",
                         kukaFeedbackRobotMpsLocked => "kukaFeedbackRobotMpsLocked",
                         kukaFeedbackRobotMpsCoupled => "kukaFeedbackRobotMpsCoupled",
                         kukaFeedbackMpsCtrlAirPressureOk => "kukaFeedbackRobotMpsCtrlAirPressureOk",
                         kukaFeedbackDockToolInPosition => "kukaFeedbackDockToolMarkerInPosition");
END_REGION
END_FUNCTION_BLOCK

FUNCTION_BLOCK "ToolInRobot"   // FB15, LAD
{ S7_Optimized_Access := 'TRUE' }
VERSION : 0.1
   VAR_INPUT
      toolIdProxy1 : Bool;
      toolIdProxy2 : Bool;
      toolIdProxy3 : Bool;
      toolIdProxy4 : Bool;
   END_VAR
   VAR_OUTPUT
      kukaFeedBackToolInRobot : Word;
      toolInRobot_Num : UInt;
   END_VAR
   VAR_TEMP
      mask : Byte;
   END_VAR
BEGIN

REGION Network 1 (SCL)

   #mask := 0;
   IF #toolIdProxy1 THEN
       #mask := #mask + 1;
   END_IF;   // bit0
   IF #toolIdProxy2 THEN
       #mask := #mask + 2;
   END_IF;   // bit1
   IF #toolIdProxy3 THEN
       #mask := #mask + 4;
   END_IF;   // bit2
   IF #toolIdProxy4 THEN
       #mask := #mask + 8;
   END_IF;   // bit3

   //Stand 1 - Tool 1 - Fork 
   //Stand 2 - Tool 2 - Pepa
   //Stand 3 - TOOL 3 - Marker
   //Stand 4 - Tool 4 - Gocator
   //Stand 5 - Tool 5 - Pole
   //Falta ajustar los sensores para que generen esas combinaciones.

   CASE #mask OF

       0:
           #toolInRobot_Num := 0;   // sin herramienta
           #kukaFeedBackToolInRobot := SWAP(UINT_TO_WORD(#toolInRobot_Num));
       1:
           #toolInRobot_Num := 2;   // PEPA
           #kukaFeedBackToolInRobot := SWAP(UINT_TO_WORD(#toolInRobot_Num));
       2:
           #toolInRobot_Num := 5;   // pole
           #kukaFeedBackToolInRobot := SWAP(UINT_TO_WORD(#toolInRobot_Num));
       3:
           #toolInRobot_Num := 1;   // fork
           #kukaFeedBackToolInRobot := SWAP(UINT_TO_WORD(#toolInRobot_Num));
          // #kukaFeedBackToolInRobot := UINT_TO_WORD(#toolInRobot_Num);  // SIN SWAP
       4:
           #toolInRobot_Num := 4;   // teaching
           #kukaFeedBackToolInRobot := SWAP(UINT_TO_WORD(#toolInRobot_Num));
       5:
           #toolInRobot_Num := 3;   // marker
           #kukaFeedBackToolInRobot := SWAP(UINT_TO_WORD(#toolInRobot_Num));
       ELSE
           #toolInRobot_Num := -1;      // combinación no válida / desconocida
   END_CASE;
END_REGION
END_FUNCTION_BLOCK

// folder: 30. Safety

FUNCTION_BLOCK "MainSafety"   // FB1, F_LAD
{ S7_Optimized_Access := 'TRUE' }
// // Functionality: Monitoring of the protective door position, light curtain and emergency stop
   VAR
      ACK_GL_Instance : ACK_GL;
      instEStopGroup : "EStopGroup";
      instLightCurtainGroup : "LightCurtainGroup";
      instSafetyDoor : "SafetyDoor";
      SafetyRobot_Instance : "SafetyRobot";
   END_VAR
   VAR_TEMP
      tempEStop1Released : Bool;
      tempEStop2Released : Bool;
      tempEStop3Released : Bool;
      tempEStop4Released : Bool;
      tempEStop5Released : Bool;
      tempEStop6Released : Bool;
      tempEStop7Released : Bool;
      tempEStop8Released : Bool;
      tempEStopAllReleased : Bool;
      tempEStopReleasedActuator : Bool;
      tempEStopAckReq : Bool;
      tempLc1Free : Bool;
      tempLc2Free : Bool;
      tempLc3Free : Bool;
      tempLc4Free : Bool;
      tempLc5Free : Bool;
      tempLc6Free : Bool;
      tempLcAllFree : Bool;
      tempLcAccessGrantedZ1 : Bool;
      tempLcAccessGrantedZ2 : Bool;
      tempLcAccessGrantedZ3 : Bool;
   END_VAR
BEGIN

REGION Network 1
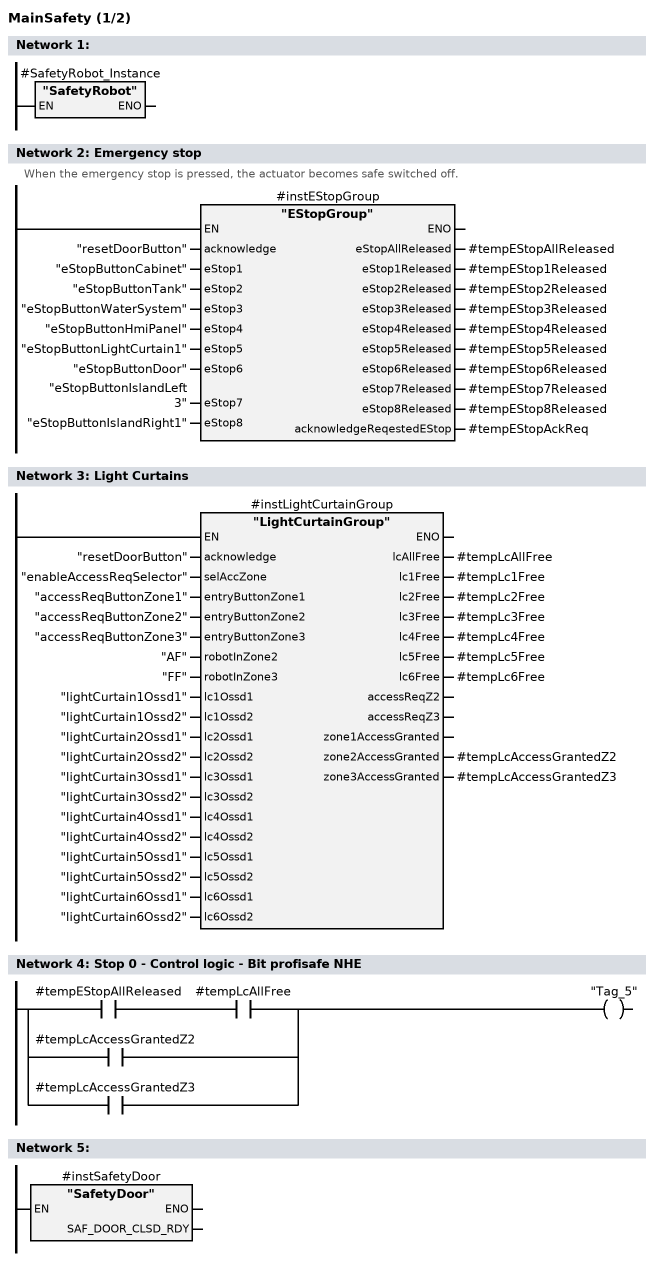
   RUNG wire#powerrail
      #SafetyRobot_Instance()
   END_RUNG
   // the same network as SCL:
   #SafetyRobot_Instance();   // "SafetyRobot"
END_REGION

REGION Network 2: Emergency stop
   // When the emergency stop is pressed, the actuator becomes safe switched off.
   RUNG wire#powerrail
      #instEStopGroup(acknowledge := "resetDoorButton", eStop1 := "eStopButtonCabinet", eStop2 := "eStopButtonTank", eStop3 := "eStopButtonWaterSystem", eStop4 := "eStopButtonHmiPanel", eStop5 := "eStopButtonLightCurtain1", eStop6 := "eStopButtonDoor", eStop7 := "eStopButtonIslandLeft 3", eStop8 := "eStopButtonIslandRight1", eStopAllReleased => #tempEStopAllReleased, eStop1Released => #tempEStop1Released, eStop2Released => #tempEStop2Released, eStop3Released => #tempEStop3Released, eStop4Released => #tempEStop4Released, eStop5Released => #tempEStop5Released, eStop6Released => #tempEStop6Released, eStop7Released => #tempEStop7Released, eStop8Released => #tempEStop8Released, acknowledgeReqestedEStop => #tempEStopAckReq)
   END_RUNG
   // the same network as SCL:
   #instEStopGroup(acknowledge := "resetDoorButton",   // "EStopGroup"
                   eStop1 := "eStopButtonCabinet",
                   eStop2 := "eStopButtonTank",
                   eStop3 := "eStopButtonWaterSystem",
                   eStop4 := "eStopButtonHmiPanel",
                   eStop5 := "eStopButtonLightCurtain1",
                   eStop6 := "eStopButtonDoor",
                   eStop7 := "eStopButtonIslandLeft 3",
                   eStop8 := "eStopButtonIslandRight1",
                   eStopAllReleased => #tempEStopAllReleased,
                   eStop1Released => #tempEStop1Released,
                   eStop2Released => #tempEStop2Released,
                   eStop3Released => #tempEStop3Released,
                   eStop4Released => #tempEStop4Released,
                   eStop5Released => #tempEStop5Released,
                   eStop6Released => #tempEStop6Released,
                   eStop7Released => #tempEStop7Released,
                   eStop8Released => #tempEStop8Released,
                   acknowledgeReqestedEStop => #tempEStopAckReq);
END_REGION

REGION Network 3: Light Curtains
   RUNG wire#powerrail
      #instLightCurtainGroup(acknowledge := "resetDoorButton", selAccZone := "enableAccessReqSelector", entryButtonZone1 := "accessReqButtonZone1", entryButtonZone2 := "accessReqButtonZone2", entryButtonZone3 := "accessReqButtonZone3", robotInZone2 := "AF", robotInZone3 := "FF", lc1Ossd1 := "lightCurtain1Ossd1", lc1Ossd2 := "lightCurtain1Ossd2", lc2Ossd1 := "lightCurtain2Ossd1", lc2Ossd2 := "lightCurtain2Ossd2", lc3Ossd1 := "lightCurtain3Ossd1", lc3Ossd2 := "lightCurtain3Ossd2", lc4Ossd1 := "lightCurtain4Ossd1", lc4Ossd2 := "lightCurtain4Ossd2", lc5Ossd1 := "lightCurtain5Ossd1", lc5Ossd2 := "lightCurtain5Ossd2", lc6Ossd1 := "lightCurtain6Ossd1", lc6Ossd2 := "lightCurtain6Ossd2", lcAllFree => #tempLcAllFree, lc1Free => #tempLc1Free, lc2Free => #tempLc2Free, lc3Free => #tempLc3Free, lc4Free => #tempLc4Free, lc5Free => #tempLc5Free, lc6Free => #tempLc6Free, accessReqZ2 =>, accessReqZ3 =>, zone1AccessGranted =>, zone2AccessGranted => #tempLcAccessGrantedZ2, zone3AccessGranted => #tempLcAccessGrantedZ3)
   END_RUNG
   // the same network as SCL:
   #instLightCurtainGroup(acknowledge := "resetDoorButton",   // "LightCurtainGroup"
                          selAccZone := "enableAccessReqSelector",
                          entryButtonZone1 := "accessReqButtonZone1",
                          entryButtonZone2 := "accessReqButtonZone2",
                          entryButtonZone3 := "accessReqButtonZone3",
                          robotInZone2 := "AF",
                          robotInZone3 := "FF",
                          lc1Ossd1 := "lightCurtain1Ossd1",
                          lc1Ossd2 := "lightCurtain1Ossd2",
                          lc2Ossd1 := "lightCurtain2Ossd1",
                          lc2Ossd2 := "lightCurtain2Ossd2",
                          lc3Ossd1 := "lightCurtain3Ossd1",
                          lc3Ossd2 := "lightCurtain3Ossd2",
                          lc4Ossd1 := "lightCurtain4Ossd1",
                          lc4Ossd2 := "lightCurtain4Ossd2",
                          lc5Ossd1 := "lightCurtain5Ossd1",
                          lc5Ossd2 := "lightCurtain5Ossd2",
                          lc6Ossd1 := "lightCurtain6Ossd1",
                          lc6Ossd2 := "lightCurtain6Ossd2",
                          lcAllFree => #tempLcAllFree,
                          lc1Free => #tempLc1Free,
                          lc2Free => #tempLc2Free,
                          lc3Free => #tempLc3Free,
                          lc4Free => #tempLc4Free,
                          lc5Free => #tempLc5Free,
                          lc6Free => #tempLc6Free,
                          zone2AccessGranted => #tempLcAccessGrantedZ2,
                          zone3AccessGranted => #tempLcAccessGrantedZ3);
END_REGION

